'~Spare FB2[273].28'; 8765 '~Spare FB2[273].29'; 8766 '~Spare FB2[273].30'; 8767 '~Spare FB2[273].31'; 8768 '~Spare FB2[274].0'; 8769 '~Spare FB2[274].1'; 8770 '~Spare FB2[274].2'; 8771 '~Spare FB2[274].3'; 8772 '~Spare FB2[274].4'; 8773 '~Spare FB2[274].5'; 8774 '~Spare FB2[274].6'; 8775 '~Spare FB2[274].7'; 8776 '~Spare FB2[274].8'; 8777 '~Spare FB2[274].9'; 8778 '~Spare FB2[274].10'; 8779 '~Spare FB2[274].11'; 8780 '~Spare FB2[274].12'; 8781 '~Spare FB2[274].13'; 8782 '~Spare FB2[274].14'; 8783 '~Spare FB2[274].15'; 8784 '~Spare FB2[274].16'; 8785 '~Spare FB2[274].17'; 8786 '~Spare FB2[274].18'; 8787 '~Spare FB2[274].19'; 8788 '~Spare FB2[274].20'; 8789 '~Spare FB2[274].21'; 8790 '~Spare FB2[274].22'; 8791 '~Spare FB2[274].23'; 8792 '~Spare FB2[274].24'; 8793 '~Spare FB2[274].25'; 8794 '~Spare FB2[274].26'; 8795 '~Spare FB2[274].27'; 8796 '~Spare FB2[274].28'; 8797 '~Spare FB2[274].29'; 8798 '~Spare FB2[274].30'; 8799 '~Spare FB2[274].31'; 8800 '~Spare FB2[275].0'; 8801 '~Spare FB2[275].1'; 8802 '~Spare FB2[275].2'; 8803 '~Spare FB2[275].3'; 8804 '~Spare FB2[275].4'; 8805 '~Spare FB2[275].5'; 8806 '~Spare FB2[275].6'; 8807 '~Spare FB2[275].7'; 8808 '~Spare FB2[275].8'; 8809 '~Spare FB2[275].9'; 8810 '~Spare FB2[275].10'; 8811 '~Spare FB2[275].11'; 8812 '~Spare FB2[275].12'; 8813 '~Spare FB2[275].13'; 8814 '~Spare FB2[275].14'; 8815 '~Spare FB2[275].15'; 8816 '~Spare FB2[275].16'; 8817 '~Spare FB2[275].17'; 8818 '~Spare FB2[275].18'; 8819 '~Spare FB2[275].19'; 8820 '~Spare FB2[275].20'; 8821 '~Spare FB2[275].21'; 8822 '~Spare FB2[275].22'; 8823 '~Spare FB2[275].23'; 8824 '~Spare FB2[275].24'; 8825 '~Spare FB2[275].25'; 8826 '~Spare FB2[275].26'; 8827 '~Spare FB2[275].27'; 8828 '~Spare FB2[275].28'; 8829 '~Spare FB2[275].29'; 8830 '~Spare FB2[275].30'; 8831 '~Spare FB2[275].31'; 8832 '~S001R13CN.I.RbtCtrlFlt - Control Fault FB2[276].0'; 8833 '~S001R13CN.I.CollDetect - Collision Detect FB2[276].1'; 8834 '~S001R13CN.Ix.RbtPromptBox - View Prompt Box at Teach Pendant FB2[276].2'; 8835 '~Spare FB2[276].3'; 8836 '~Spare FB2[276].4'; 8837 '~Spare FB2[276].5'; 8838 '~Spare FB2[276].6'; 8839 '~Spare FB2[276].7'; 8840 '~Spare FB2[276].8'; 8841 '~Spare FB2[276].9'; 8842 '~Spare FB2[276].10'; 8843 '~S001R13CN.I.Wc1WldFlt -Weld Controller 1 Weld Fault FB2[276].11'; 8844 '~S001R13CN.I.Wc1Flt - Weld Timer Flt - Depress Man Weld To Continue FB2[276].12'; 8845 '~S001R13CN.I.Wc1SGunFlt - Weld Controller 1 Servo Gun Fault FB2[276].13'; 8846 '~S001R13CN.I.Wc1SGunMtrTempFlt - Cntrl 1 Servo Gun Motor Over Temp FB2[276].14'; 8847 '~S001R13CN.I.Td1MtrFlt - Tip Dress 1 Motor Fault FB2[276].15'; 8848 '~S001R13CN.I.WC1XfmrTempFlt - Weld Cntrl 1 Transformer Over Temp FB2[276].16'; 8849 '~S001R13CN.I.AutoTipChng1Flt - Auto Tip Changer 1 Fault FB2[276].17'; 8850 '~S001R13CN.I.Slr1NotReady - Seal Controller 1 Not Ready FB2[276].18'; 8851 '~S001R13CN.I.Slr1MajorFlt - Seal Controller 1 Major Fault FB2[276].19'; 8852 '~S001R13CN.I.Slr1VolNotOk - Seal Controller 1 Volume Not Ok Fault FB2[276].20'; 8853 '~S001R13CN.I.Slr1PurgeFlt - Seal Controller 1 Purge Fault FB2[276].21'; 8854 '~S001R13CN.I.Slr1DoserNot Filled - Seal Cntrl 1 Doser Not Filled FB2[276].22'; 8855 '~S001R13CN.I.Slr1No2ClnMxr - Seal Cntrl1 No 2C In Mixer Fault FB2[276].23'; 8856 '~S001R13CN.I.Slr1NzlBroken - Seal Controller 1 Nozzle Broken Fault FB2[276].24'; 8857 '~S001R13CN.I.Slr1NozzleChgReq - Seal Cntrl1 Nozzle Change Reqd FB2[276].25'; 8858 '~S001R13CN.I.Slr1CycleInterrupted - Seal Cntrl1 Cycle Interrupted FB2[276].26'; 8859 '~S001R13CN.I.Stdw1Flt - Stud Weld 1 Weld Fault FB2[276].27'; 8860 '~S001R13CN.I.Stdw1DlyExcdd - Stud Weld 1 Time Delay Exceeded Flt FB2[276].28'; 8861 '~S001R13CN.I.Stdw1Maint Reqd - Stud Weld 1 Maintenance Required FB2[276].29'; 8862 '~S001R13CN.I.Stdw1Reject - Stud Weld 1 art Reject Fault FB2[276].30'; 8863 '~S001R13CN.I.Rvt1Flt - Rivet Controller 1 Fault FB2[276].31'; 8864 '~S001R13CN.I.Rvt1DlyExcdd - Rivet Cntrl 1 Time Delay Exceeded Flt FB2[277].0'; 8865 '~S001R13CN.I.AutoPulledTipByp1 - Auto Pulled Tip Bypass 1 FB2[277].1'; 8866 '~S001R13CN.I.StdWld1EquipmentFlt - Stud Weld 1 Equipment Fault FB2[277].2'; 8867 '~S001R13CN.I.StdWld1BrcktNotPresent - Stud Weld 1 Bracket Not Pres FB2[277].3'; 8868 '~S001R13CN.I.PierceFlt - Pierce Fault FB2[277].4'; 8869 '~S001R13CN.I.NoVisionMeasErr - Vision System Measurement Error FB2[277].5'; 8870 '~S001R13CN.I.VisionSysCalErr - Vision System Calibration Fault FB2[277].6'; 8871 '~S001R13CN.I.VisionSysErr - Vision System Error FB2[277].7'; 8872 '~S001R13CN.I.RackOutOfTolerance - Vision Sys Rack Out Of Tolerance FB2[277].8'; 8873 '~S001R13CN.Ix.TorqFlt - Torque Not Ok FB2[277].9'; 8874 '~S001R13CN.Ix.MwFlt - Mig Weld Controller Fault FB2[277].10'; 8875 '~S001R13CN.Ix.MwWireStuckFlt - Mig Welder Wire Stuck FB2[277].11'; 8876 '~S001R13CN.Ix.MwWldFlt - Mig Welder Bad Bronze Weld Indicator Flt FB2[277].12'; 8877 '~S001R13CN.I.O.TipChngReqd1 - Weld Cntrl 1 Tip Change Required FB2[277].13'; 8878 '~S001R13CN.I.M.NutDetectFlt1 - Nut Welder 1 Nut Detection Fault FB2[277].14'; 8879 '~S001R13CN.I.M.NutProjFlt1 - Nut Welder 1 Weld Not In Tolerance FB2[277].15'; 8880 '~S001R13CN.M.WrongRivetAtNose - Remove Wrong Rivet At Nose FB2[277].16'; 8881 '~S001R13CN.Ix.MwWldLimitErr - Mig Welder CurrentVoltage Out of Tolerance FB2[277].17'; 8882 '~S001R13CN.Ix.MigRdy Mig Welder Not Ready FB2[277].18'; 8883 '~Spare FB2[277].19'; 8884 '~Spare FB2[277].20'; 8885 '~S001R13CN.I.Wc2WldFlt -Weld Controller 2 Weld Fault FB2[277].21'; 8886 '~S001R13CN.I.Wc2Flt - Weld Timer Flt - Depress Man Weld To Continue FB2[277].22'; 8887 '~S001R13CN.I.Wc2SGunFlt - Weld Controller 2 Servo Gun Fault FB2[277].23'; 8888 '~S001R13CN.I.Wc2SGunMtrTempFlt - Cntrl 2 Servo Gun Motor Over Temp FB2[277].24'; 8889 '~S001R13CN.I.Td2MtrFlt - Tip Dress 2 Motor Fault FB2[277].25'; 8890 '~S001R13CN.I.WC2XfmrTempFlt - Weld Cntrl 2 Transformer Over Temp FB2[277].26'; 8891 '~S001R13CN.I.AutoTipChng2Flt - Auto Tip Changer 2 Fault FB2[277].27'; 8892 '~S001R13CN.I.Slr2NotReady - Seal Controller 2 Not Ready FB2[277].28'; 8893 '~S001R13CN.I.Slr2MajorFlt - Seal Controller 2 Major Fault FB2[277].29'; 8894 '~S001R13CN.I.Slr2VolNotOk - Seal Controller 2 Volume Not Ok Fault FB2[277].30'; 8895 '~S001R13CN.I.Slr2PurgeFlt - Seal Controller 2 Purge Fault FB2[277].31'; 8896 '~S001R13CN.I.Slr2DoserNot Filled - Seal Cntrl 2 Doser Not Filled FB2[278].0'; 8897 '~S001R13CN.I.Slr2No2ClnMxr - Seal Cntrl2 No 2C In Mixer Fault FB2[278].1'; 8898 '~S001R13CN.I.Slr2NzlBroken - Seal Controller 2 Nozzle Broken Fault FB2[278].2'; 8899 '~S001R13CN.I.Slr2NozzleChgReq - Seal Cntrl2 Nozzle Change Reqd FB2[278].3'; 8900 '~S001R13CN.I.Slr2CycleInterrupted - Seal Cntrl2 Cycle Interrupted FB2[278].4'; 8901 '~S001R13CN.I.Stdw2Flt - Stud Weld 2 Weld Fault FB2[278].5'; 8902 '~S001R13CN.I.Stdw2DlyExcdd - Stud Weld 2 Time Delay Exceeded Flt FB2[278].6'; 8903 '~S001R13CN.I.Stdw2Maint Reqd - Stud Weld 2 Maintenance Required FB2[278].7'; 8904 '~S001R13CN.I.Stdw2Reject - Stud Weld 2 art Reject Fault FB2[278].8'; 8905 '~S001R13CN.I.Rvt2Flt - Rivet Controller 2 Fault FB2[278].9'; 8906 '~S001R13CN.I.Rvt2DlyExcdd - Rivet Cntrl 2 Time Delay Exceeded Flt FB2[278].10'; 8907 '~S001R13CN.I.AutoPulledTipByp2 - Auto Pulled Tip Bypass 2 FB2[278].11'; 8908 '~S001R13CN.I.StdWld2EquipmentFlt - Stud Weld 2 Equipment Fault FB2[278].12'; 8909 '~S001R13CN.I.StdWld2BrcktNotPresent - Stud Weld 2 Bracket Not Pres FB2[278].13'; 8910 '~S001R13CN.Ix.LsrWldMntrFlt - Seam Geometry/Laser Weld Monitor Flt FB2[278].14'; 8911 '~S001R13CN.Ix.LsrHeadFlt - Laser Head Fault FB2[278].15'; 8912 '~S001R13CN.Ix.LsrGlsFlt - Glass Fault FB2[278].16'; 8913 '~S001R13CN.Ix.LsrWhlFlt - Pressure Wheel Not In Range Fault FB2[278].17'; 8914 '~S001R13CN.Ix.LsrGeoFlt - Seam Geometry/Laser Bad Process Geo Flt FB2[278].18'; 8915 '~S001R13CN.Ix.LsrHdCollFlt - Laser Head Collision Fault FB2[278].19'; 8916 '~S001R13CN.Ix.LsrHdSysFlt - Laser Head System Fault FB2[278].20'; 8917 '~S001R13CN.Ix.LsrHdFar - Laser Head Far Fault FB2[278].21'; 8918 '~S001R13CN.Ix.LsrHdSftCollFlt - Laser Head Software Collision Flt FB2[278].22'; 8919 '~S001R13CN.I.O.TipChngReqd2 - Weld Cntrl 2 Tip Change Required FB2[278].23'; 8920 '~S001R13CN.I.M.NutDetectFlt2 - Nut Welder 2 Nut Detection Fault FB2[278].24'; 8921 '~S001R13CN.I.M.NutProjFlt2 - Nut Welder 2 Weld Not In Tolerance FB2[278].25'; 8922 '~S001R13CN.I.TCWrongToolInStand - Tool Changer Wrong Tool In Stand FB2[278].26'; 8923 '~Spare FB2[278].27'; 8924 '~Spare FB2[278].28'; 8925 '~Spare FB2[278].29'; 8926 '~Spare FB2[278].30'; 8927 '~Spare FB2[278].31'; 8928 '~S001R13CN.I.VisionCommOK - Vision System Comm Fault FB2[279].0'; 8929 '~S001R13CN.I.OutOfTolerance - Vision System Out Of Tolerance FB2[279].1'; 8930 '~S001R13CN.I.MeasureReject - Vision System Measure Reject FB2[279].2'; 8931 '~S001R13CN.I.VisionSysCalibrationFlt - Vision System Calibration Flt FB2[279].3'; 8932 '~S001R13CN.I.VisionSysFlt - Vision System Flt FB2[279].4'; 8933 '~Spare FB2[279].5'; 8934 '~Spare FB2[279].6'; 8935 '~Spare FB2[279].7'; 8936 '~Spare FB2[279].8'; 8937 '~Spare FB2[279].9'; 8938 '~Spare FB2[279].10'; 8939 '~Spare FB2[279].11'; 8940 '~Spare FB2[279].12'; 8941 '~Spare FB2[279].13'; 8942 '~Spare FB2[279].14'; 8943 '~Spare FB2[279].15'; 8944 '~Spare FB2[279].16'; 8945 '~Spare FB2[279].17'; 8946 '~S001R13CN.M.InteruptCyc - Laser Cyc Interupt Cut Wire And Reject Car FB2[279].18'; 8947 '~S001R13CN.M.SuspectPart Inspect Vehicle And Accept Or Reject FB2[279].19'; 8948 '~S001R13 Power Meter High Power Fault Detected FB2[279].20'; 8949 '~S001R13 Power Meter Low Power Fault Detected FB2[279].21'; 8950 '~Spare FB2[279].22'; 8951 '~Spare FB2[279].23'; 8952 '~Spare FB2[279].24'; 8953 '~Spare FB2[279].25'; 8954 '~Spare FB2[279].26'; 8955 '~Spare FB2[279].27'; 8956 '~Spare FB2[279].28'; 8957 '~Spare FB2[279].29'; 8958 '~Spare FB2[279].30'; 8959 '~Spare FB2[279].31'; 8960 '~Spare FB2[280].0'; 8961 '~Spare FB2[280].1'; 8962 '~Spare FB2[280].2'; 8963 '~Spare FB2[280].3'; 8964 '~Spare FB2[280].4'; 8965 '~Spare FB2[280].5'; 8966 '~Spare FB2[280].6'; 8967 '~Spare FB2[280].7'; 8968 '~Spare FB2[280].8'; 8969 '~Spare FB2[280].9'; 8970 '~Spare FB2[280].10'; 8971 '~Spare FB2[280].11'; 8972 '~Spare FB2[280].12'; 8973 '~Spare FB2[280].13'; 8974 '~Spare FB2[280].14'; 8975 '~Spare FB2[280].15'; 8976 '~Spare FB2[280].16'; 8977 '~Spare FB2[280].17'; 8978 '~Spare FB2[280].18'; 8979 '~Spare FB2[280].19'; 8980 '~Spare FB2[280].20'; 8981 '~Spare FB2[280].21'; 8982 '~Spare FB2[280].22'; 8983 '~Spare FB2[280].23'; 8984 '~Spare FB2[280].24'; 8985 '~Spare FB2[280].25'; 8986 '~Spare FB2[280].26'; 8987 '~Spare FB2[280].27'; 8988 '~Spare FB2[280].28'; 8989 '~Spare FB2[280].29'; 8990 '~Spare FB2[280].30'; 8991 '~Spare FB2[280].31'; 8992 '~Spare FB2[281].0'; 8993 '~Spare FB2[281].1'; 8994 '~Spare FB2[281].2'; 8995 '~Spare FB2[281].3'; 8996 '~Spare FB2[281].4'; 8997 '~Spare FB2[281].5'; 8998 '~Spare FB2[281].6'; 8999 '~Spare FB2[281].7'; 9000 '~Spare FB2[281].8'; 9001 '~Spare FB2[281].9'; 9002 '~Spare FB2[281].10'; 9003 '~Spare FB2[281].11'; 9004 '~Spare FB2[281].12'; 9005 '~Spare FB2[281].13'; 9006 '~Spare FB2[281].14'; 9007 '~Spare FB2[281].15'; 9008 '~Spare FB2[281].16'; 9009 '~Spare FB2[281].17'; 9010 '~Spare FB2[281].18'; 9011 '~Spare FB2[281].19'; 9012 '~Spare FB2[281].20'; 9013 '~Spare FB2[281].21'; 9014 '~Spare FB2[281].22'; 9015 '~Spare FB2[281].23'; 9016 '~Spare FB2[281].24'; 9017 '~Spare FB2[281].25'; 9018 '~Spare FB2[281].26'; 9019 '~Spare FB2[281].27'; 9020 '~Spare FB2[281].28'; 9021 '~Spare FB2[281].29'; 9022 '~Spare FB2[281].30'; 9023 '~Spare FB2[281].31'; 9024 '~Spare FB2[282].0'; 9025 '~Spare FB2[282].1'; 9026 '~Spare FB2[282].2'; 9027 '~Spare FB2[282].3'; 9028 '~Spare FB2[282].4'; 9029 '~Spare FB2[282].5'; 9030 '~Spare FB2[282].6'; 9031 '~Spare FB2[282].7'; 9032 '~Spare FB2[282].8'; 9033 '~Spare FB2[282].9'; 9034 '~Spare FB2[282].10'; 9035 '~Spare FB2[282].11'; 9036 '~Spare FB2[282].12'; 9037 '~Spare FB2[282].13'; 9038 '~Spare FB2[282].14'; 9039 '~Spare FB2[282].15'; 9040 '~Spare FB2[282].16'; 9041 '~Spare FB2[282].17'; 9042 '~Spare FB2[282].18'; 9043 '~Spare FB2[282].19'; 9044 '~Spare FB2[282].20'; 9045 '~Spare FB2[282].21'; 9046 '~Spare FB2[282].22'; 9047 '~Spare FB2[282].23'; 9048 '~Spare FB2[282].24'; 9049 '~Spare FB2[282].25'; 9050 '~Spare FB2[282].26'; 9051 '~Spare FB2[282].27'; 9052 '~Spare FB2[282].28'; 9053 '~Spare FB2[282].29'; 9054 '~Spare FB2[282].30'; 9055 '~Spare FB2[282].31'; 9056 '~Spare FB2[283].0'; 9057 '~Spare FB2[283].1'; 9058 '~Spare FB2[283].2'; 9059 '~Spare FB2[283].3'; 9060 '~Spare FB2[283].4'; 9061 '~Spare FB2[283].5'; 9062 '~Spare FB2[283].6'; 9063 '~Spare FB2[283].7'; 9064 '~Spare FB2[283].8'; 9065 '~Spare FB2[283].9'; 9066 '~Spare FB2[283].10'; 9067 '~Spare FB2[283].11'; 9068 '~Spare FB2[283].12'; 9069 '~Spare FB2[283].13'; 9070 '~Spare FB2[283].14'; 9071 '~Spare FB2[283].15'; 9072 '~Spare FB2[283].16'; 9073 '~Spare FB2[283].17'; 9074 '~Spare FB2[283].18'; 9075 '~Spare FB2[283].19'; 9076 '~Spare FB2[283].20'; 9077 '~Spare FB2[283].21'; 9078 '~Spare FB2[283].22'; 9079 '~Spare FB2[283].23'; 9080 '~Spare FB2[283].24'; 9081 '~Spare FB2[283].25'; 9082 '~Spare FB2[283].26'; 9083 '~Spare FB2[283].27'; 9084 '~Spare FB2[283].28'; 9085 '~Spare FB2[283].29'; 9086 '~Spare FB2[283].30'; 9087 '~Spare FB2[283].31'; 9088 '~S001R14CN.I.RbtCtrlFlt - Control Fault FB2[284].0'; 9089 '~S001R14CN.I.CollDetect - Collision Detect FB2[284].1'; 9090 '~S001R14CN.Ix.RbtPromptBox - View Prompt Box at Teach Pendant FB2[284].2'; 9091 '~Spare FB2[284].3'; 9092 '~Spare FB2[284].4'; 9093 '~Spare FB2[284].5'; 9094 '~Spare FB2[284].6'; 9095 '~Spare FB2[284].7'; 9096 '~Spare FB2[284].8'; 9097 '~Spare FB2[284].9'; 9098 '~Spare FB2[284].10'; 9099 '~S001R14CN.I.Wc1WldFlt -Weld Controller 1 Weld Fault FB2[284].11'; 9100 '~S001R14CN.I.Wc1Flt - Weld Timer Flt - Depress Man Weld To Continue FB2[284].12'; 9101 '~S001R14CN.I.Wc1SGunFlt - Weld Controller 1 Servo Gun Fault FB2[284].13'; 9102 '~S001R14CN.I.Wc1SGunMtrTempFlt - Cntrl 1 Servo Gun Motor Over Temp FB2[284].14'; 9103 '~S001R14CN.I.Td1MtrFlt - Tip Dress 1 Motor Fault FB2[284].15'; 9104 '~S001R14CN.I.WC1XfmrTempFlt - Weld Cntrl 1 Transformer Over Temp FB2[284].16'; 9105 '~S001R14CN.I.AutoTipChng1Flt - Auto Tip Changer 1 Fault FB2[284].17'; 9106 '~S001R14CN.I.Slr1NotReady - Seal Controller 1 Not Ready FB2[284].18'; 9107 '~S001R14CN.I.Slr1MajorFlt - Seal Controller 1 Major Fault FB2[284].19'; 9108 '~S001R14CN.I.Slr1VolNotOk - Seal Controller 1 Volume Not Ok Fault FB2[284].20'; 9109 '~S001R14CN.I.Slr1PurgeFlt - Seal Controller 1 Purge Fault FB2[284].21'; 9110 '~S001R14CN.I.Slr1DoserNot Filled - Seal Cntrl 1 Doser Not Filled FB2[284].22'; 9111 '~S001R14CN.I.Slr1No2ClnMxr - Seal Cntrl1 No 2C In Mixer Fault FB2[284].23'; 9112 '~S001R14CN.I.Slr1NzlBroken - Seal Controller 1 Nozzle Broken Fault FB2[284].24'; 9113 '~S001R14CN.I.Slr1NozzleChgReq - Seal Cntrl1 Nozzle Change Reqd FB2[284].25'; 9114 '~S001R14CN.I.Slr1CycleInterrupted - Seal Cntrl1 Cycle Interrupted FB2[284].26'; 9115 '~S001R14CN.I.Stdw1Flt - Stud Weld 1 Weld Fault FB2[284].27'; 9116 '~S001R14CN.I.Stdw1DlyExcdd - Stud Weld 1 Time Delay Exceeded Flt FB2[284].28'; 9117 '~S001R14CN.I.Stdw1Maint Reqd - Stud Weld 1 Maintenance Required FB2[284].29'; 9118 '~S001R14CN.I.Stdw1Reject - Stud Weld 1 art Reject Fault FB2[284].30'; 9119 '~S001R14CN.I.Rvt1Flt - Rivet Controller 1 Fault FB2[284].31'; 9120 '~S001R14CN.I.Rvt1DlyExcdd - Rivet Cntrl 1 Time Delay Exceeded Flt FB2[285].0'; 9121 '~S001R14CN.I.AutoPulledTipByp1 - Auto Pulled Tip Bypass 1 FB2[285].1'; 9122 '~S001R14CN.I.StdWld1EquipmentFlt - Stud Weld 1 Equipment Fault FB2[285].2'; 9123 '~S001R14CN.I.StdWld1BrcktNotPresent - Stud Weld 1 Bracket Not Pres FB2[285].3'; 9124 '~S001R14CN.I.PierceFlt - Pierce Fault FB2[285].4'; 9125 '~S001R14CN.I.NoVisionMeasErr - Vision System Measurement Error FB2[285].5'; 9126 '~S001R14CN.I.VisionSysCalErr - Vision System Calibration Fault FB2[285].6'; 9127 '~S001R14CN.I.VisionSysErr - Vision System Error FB2[285].7'; 9128 '~S001R14CN.I.RackOutOfTolerance - Vision Sys Rack Out Of Tolerance FB2[285].8'; 9129 '~S001R14CN.Ix.TorqFlt - Torque Not Ok FB2[285].9'; 9130 '~S001R14CN.Ix.MwFlt - Mig Weld Controller Fault FB2[285].10'; 9131 '~S001R14CN.Ix.MwWireStuckFlt - Mig Welder Wire Stuck FB2[285].11'; 9132 '~S001R14CN.Ix.MwWldFlt - Mig Welder Bad Bronze Weld Indicator Flt FB2[285].12'; 9133 '~S001R14CN.I.O.TipChngReqd1 - Weld Cntrl 1 Tip Change Required FB2[285].13'; 9134 '~S001R14CN.I.M.NutDetectFlt1 - Nut Welder 1 Nut Detection Fault FB2[285].14'; 9135 '~S001R14CN.I.M.NutProjFlt1 - Nut Welder 1 Weld Not In Tolerance FB2[285].15'; 9136 '~S001R14CN.M.WrongRivetAtNose - Remove Wrong Rivet At Nose FB2[285].16'; 9137 '~S001R14CN.Ix.MwWldLimitErr - Mig Welder CurrentVoltage Out of Tolerance FB2[285].17'; 9138 '~S001R14CN.Ix.MigRdy Mig Welder Not Ready FB2[285].18'; 9139 '~Spare FB2[285].19'; 9140 '~Spare FB2[285].20'; 9141 '~S001R14CN.I.Wc2WldFlt -Weld Controller 2 Weld Fault FB2[285].21'; 9142 '~S001R14CN.I.Wc2Flt - Weld Timer Flt - Depress Man Weld To Continue FB2[285].22'; 9143 '~S001R14CN.I.Wc2SGunFlt - Weld Controller 2 Servo Gun Fault FB2[285].23'; 9144 '~S001R14CN.I.Wc2SGunMtrTempFlt - Cntrl 2 Servo Gun Motor Over Temp FB2[285].24'; 9145 '~S001R14CN.I.Td2MtrFlt - Tip Dress 2 Motor Fault FB2[285].25'; 9146 '~S001R14CN.I.WC2XfmrTempFlt - Weld Cntrl 2 Transformer Over Temp FB2[285].26'; 9147 '~S001R14CN.I.AutoTipChng2Flt - Auto Tip Changer 2 Fault FB2[285].27'; 9148 '~S001R14CN.I.Slr2NotReady - Seal Controller 2 Not Ready FB2[285].28'; 9149 '~S001R14CN.I.Slr2MajorFlt - Seal Controller 2 Major Fault FB2[285].29'; 9150 '~S001R14CN.I.Slr2VolNotOk - Seal Controller 2 Volume Not Ok Fault FB2[285].30'; 9151 '~S001R14CN.I.Slr2PurgeFlt - Seal Controller 2 Purge Fault FB2[285].31'; 9152 '~S001R14CN.I.Slr2DoserNot Filled - Seal Cntrl 2 Doser Not Filled FB2[286].0'; 9153 '~S001R14CN.I.Slr2No2ClnMxr - Seal Cntrl2 No 2C In Mixer Fault FB2[286].1'; 9154 '~S001R14CN.I.Slr2NzlBroken - Seal Controller 2 Nozzle Broken Fault FB2[286].2'; 9155 '~S001R14CN.I.Slr2NozzleChgReq - Seal Cntrl2 Nozzle Change Reqd FB2[286].3'; 9156 '~S001R14CN.I.Slr2CycleInterrupted - Seal Cntrl2 Cycle Interrupted FB2[286].4'; 9157 '~S001R14CN.I.Stdw2Flt - Stud Weld 2 Weld Fault FB2[286].5'; 9158 '~S001R14CN.I.Stdw2DlyExcdd - Stud Weld 2 Time Delay Exceeded Flt FB2[286].6'; 9159 '~S001R14CN.I.Stdw2Maint Reqd - Stud Weld 2 Maintenance Required FB2[286].7'; 9160 '~S001R14CN.I.Stdw2Reject - Stud Weld 2 art Reject Fault FB2[286].8'; 9161 '~S001R14CN.I.Rvt2Flt - Rivet Controller 2 Fault FB2[286].9'; 9162 '~S001R14CN.I.Rvt2DlyExcdd - Rivet Cntrl 2 Time Delay Exceeded Flt FB2[286].10'; 9163 '~S001R14CN.I.AutoPulledTipByp2 - Auto Pulled Tip Bypass 2 FB2[286].11'; 9164 '~S001R14CN.I.StdWld2EquipmentFlt - Stud Weld 2 Equipment Fault FB2[286].12'; 9165 '~S001R14CN.I.StdWld2BrcktNotPresent - Stud Weld 2 Bracket Not Pres FB2[286].13'; 9166 '~S001R14CN.Ix.LsrWldMntrFlt - Seam Geometry/Laser Weld Monitor Flt FB2[286].14'; 9167 '~S001R14CN.Ix.LsrHeadFlt - Laser Head Fault FB2[286].15'; 9168 '~S001R14CN.Ix.LsrGlsFlt - Glass Fault FB2[286].16'; 9169 '~S001R14CN.Ix.LsrWhlFlt - Pressure Wheel Not In Range Fault FB2[286].17'; 9170 '~S001R14CN.Ix.LsrGeoFlt - Seam Geometry/Laser Bad Process Geo Flt FB2[286].18'; 9171 '~S001R14CN.Ix.LsrHdCollFlt - Laser Head Collision Fault FB2[286].19'; 9172 '~S001R14CN.Ix.LsrHdSysFlt - Laser Head System Fault FB2[286].20'; 9173 '~S001R14CN.Ix.LsrHdFar - Laser Head Far Fault FB2[286].21'; 9174 '~S001R14CN.Ix.LsrHdSftCollFlt - Laser Head Software Collision Flt FB2[286].22'; 9175 '~S001R14CN.I.O.TipChngReqd2 - Weld Cntrl 2 Tip Change Required FB2[286].23'; 9176 '~S001R14CN.I.M.NutDetectFlt2 - Nut Welder 2 Nut Detection Fault FB2[286].24'; 9177 '~S001R14CN.I.M.NutProjFlt2 - Nut Welder 2 Weld Not In Tolerance FB2[286].25'; 9178 '~S001R14CN.I.TCWrongToolInStand - Tool Changer Wrong Tool In Stand FB2[286].26'; 9179 '~Spare FB2[286].27'; 9180 '~Spare FB2[286].28'; 9181 '~Spare FB2[286].29'; 9182 '~Spare FB2[286].30'; 9183 '~Spare FB2[286].31'; 9184 '~S001R14CN.I.VisionCommOK - Vision System Comm Fault FB2[287].0'; 9185 '~S001R14CN.I.OutOfTolerance - Vision System Out Of Tolerance FB2[287].1'; 9186 '~S001R14CN.I.MeasureReject - Vision System Measure Reject FB2[287].2'; 9187 '~S001R14CN.I.VisionSysCalibrationFlt - Vision System Calibration Flt FB2[287].3'; 9188 '~S001R14CN.I.VisionSysFlt - Vision System Flt FB2[287].4'; 9189 '~Spare FB2[287].5'; 9190 '~Spare FB2[287].6'; 9191 '~Spare FB2[287].7'; 9192 '~Spare FB2[287].8'; 9193 '~Spare FB2[287].9'; 9194 '~Spare FB2[287].10'; 9195 '~Spare FB2[287].11'; 9196 '~Spare FB2[287].12'; 9197 '~Spare FB2[287].13'; 9198 '~Spare FB2[287].14'; 9199 '~Spare FB2[287].15'; 9200 '~Spare FB2[287].16'; 9201 '~Spare FB2[287].17'; 9202 '~S001R14CN.M.InteruptCyc - Laser Cyc Interupt Cut Wire And Reject Car FB2[287].18'; 9203 '~S001R14CN.M.SuspectPart Inspect Vehicle And Accept Or Reject FB2[287].19'; 9204 '~S001R14 Power Meter High Power Fault Detected FB2[287].20'; 9205 '~S001R14 Power Meter Low Power Fault Detected FB2[287].21'; 9206 '~Spare FB2[287].22'; 9207 '~Spare FB2[287].23'; 9208 '~Spare FB2[287].24'; 9209 '~Spare FB2[287].25'; 9210 '~Spare FB2[287].26'; 9211 '~Spare FB2[287].27'; 9212 '~Spare FB2[287].28'; 9213 '~Spare FB2[287].29'; 9214 '~Spare FB2[287].30'; 9215 '~Spare FB2[287].31'; 9216 '~Spare FB2[288].0'; 9217 '~Spare FB2[288].1'; 9218 '~Spare FB2[288].2'; 9219 '~Spare FB2[288].3'; 9220 '~Spare FB2[288].4'; 9221 '~Spare FB2[288].5'; 9222 '~Spare FB2[288].6'; 9223 '~Spare FB2[288].7'; 9224 '~Spare FB2[288].8'; 9225 '~Spare FB2[288].9'; 9226 '~Spare FB2[288].10'; 9227 '~Spare FB2[288].11'; 9228 '~Spare FB2[288].12'; 9229 '~Spare FB2[288].13'; 9230 '~Spare FB2[288].14'; 9231 '~Spare FB2[288].15'; 9232 '~Spare FB2[288].16'; 9233 '~Spare FB2[288].17'; 9234 '~Spare FB2[288].18'; 9235 '~Spare FB2[288].19'; 9236 '~Spare FB2[288].20'; 9237 '~Spare FB2[288].21'; 9238 '~Spare FB2[288].22'; 9239 '~Spare FB2[288].23'; 9240 '~Spare FB2[288].24'; 9241 '~Spare FB2[288].25'; 9242 '~Spare FB2[288].26'; 9243 '~Spare FB2[288].27'; 9244 '~Spare FB2[288].28'; 9245 '~Spare FB2[288].29'; 9246 '~Spare FB2[288].30'; 9247 '~Spare FB2[288].31'; 9248 '~Spare FB2[289].0'; 9249 '~Spare FB2[289].1'; 9250 '~Spare FB2[289].2'; 9251 '~Spare FB2[289].3'; 9252 '~Spare FB2[289].4'; 9253 '~Spare FB2[289].5'; 9254 '~Spare FB2[289].6'; 9255 '~Spare FB2[289].7'; 9256 '~Spare FB2[289].8'; 9257 '~Spare FB2[289].9'; 9258 '~Spare FB2[289].10'; 9259 '~Spare FB2[289].11'; 9260 '~Spare FB2[289].12'; 9261 '~Spare FB2[289].13'; 9262 '~Spare FB2[289].14'; 9263 '~Spare FB2[289].15'; 9264 '~Spare FB2[289].16'; 9265 '~Spare FB2[289].17'; 9266 '~Spare FB2[289].18'; 9267 '~Spare FB2[289].19'; 9268 '~Spare FB2[289].20'; 9269 '~Spare FB2[289].21'; 9270 '~Spare FB2[289].22'; 9271 '~Spare FB2[289].23'; 9272 '~Spare FB2[289].24'; 9273 '~Spare FB2[289].25'; 9274 '~Spare FB2[289].26'; 9275 '~Spare FB2[289].27'; 9276 '~Spare FB2[289].28'; 9277 '~Spare FB2[289].29'; 9278 '~Spare FB2[289].30'; 9279 '~Spare FB2[289].31'; 9280 '~Spare FB2[290].0'; 9281 '~Spare FB2[290].1'; 9282 '~Spare FB2[290].2'; 9283 '~Spare FB2[290].3'; 9284 '~Spare FB2[290].4'; 9285 '~Spare FB2[290].5'; 9286 '~Spare FB2[290].6'; 9287 '~Spare FB2[290].7'; 9288 '~Spare FB2[290].8'; 9289 '~Spare FB2[290].9'; 9290 '~Spare FB2[290].10'; 9291 '~Spare FB2[290].11'; 9292 '~Spare FB2[290].12'; 9293 '~Spare FB2[290].13'; 9294 '~Spare FB2[290].14'; 9295 '~Spare FB2[290].15'; 9296 '~Spare FB2[290].16'; 9297 '~Spare FB2[290].17'; 9298 '~Spare FB2[290].18'; 9299 '~Spare FB2[290].19'; 9300 '~Spare FB2[290].20'; 9301 '~Spare FB2[290].21'; 9302 '~Spare FB2[290].22'; 9303 '~Spare FB2[290].23'; 9304 '~Spare FB2[290].24'; 9305 '~Spare FB2[290].25'; 9306 '~Spare FB2[290].26'; 9307 '~Spare FB2[290].27'; 9308 '~Spare FB2[290].28'; 9309 '~Spare FB2[290].29'; 9310 '~Spare FB2[290].30'; 9311 '~Spare FB2[290].31'; 9312 '~Spare FB2[291].0'; 9313 '~Spare FB2[291].1'; 9314 '~Spare FB2[291].2'; 9315 '~Spare FB2[291].3'; 9316 '~Spare FB2[291].4'; 9317 '~Spare FB2[291].5'; 9318 '~Spare FB2[291].6'; 9319 '~Spare FB2[291].7'; 9320 '~Spare FB2[291].8'; 9321 '~Spare FB2[291].9'; 9322 '~Spare FB2[291].10'; 9323 '~Spare FB2[291].11'; 9324 '~Spare FB2[291].12'; 9325 '~Spare FB2[291].13'; 9326 '~Spare FB2[291].14'; 9327 '~Spare FB2[291].15'; 9328 '~Spare FB2[291].16'; 9329 '~Spare FB2[291].17'; 9330 '~Spare FB2[291].18'; 9331 '~Spare FB2[291].19'; 9332 '~Spare FB2[291].20'; 9333 '~Spare FB2[291].21'; 9334 '~Spare FB2[291].22'; 9335 '~Spare FB2[291].23'; 9336 '~Spare FB2[291].24'; 9337 '~Spare FB2[291].25'; 9338 '~Spare FB2[291].26'; 9339 '~Spare FB2[291].27'; 9340 '~Spare FB2[291].28'; 9341 '~Spare FB2[291].29'; 9342 '~Spare FB2[291].30'; 9343 '~Spare FB2[291].31'; 9344 '~S001R15CN.I.RbtCtrlFlt - Control Fault FB2[292].0'; 9345 '~S001R15CN.I.CollDetect - Collision Detect FB2[292].1'; 9346 '~S001R15CN.Ix.RbtPromptBox - View Prompt Box at Teach Pendant FB2[292].2'; 9347 '~Spare FB2[292].3'; 9348 '~Spare FB2[292].4'; 9349 '~Spare FB2[292].5'; 9350 '~Spare FB2[292].6'; 9351 '~Spare FB2[292].7'; 9352 '~Spare FB2[292].8'; 9353 '~Spare FB2[292].9'; 9354 '~Spare FB2[292].10'; 9355 '~S001R15CN.I.Wc1WldFlt -Weld Controller 1 Weld Fault FB2[292].11'; 9356 '~S001R15CN.I.Wc1Flt - Weld Timer Flt - Depress Man Weld To Continue FB2[292].12'; 9357 '~S001R15CN.I.Wc1SGunFlt - Weld Controller 1 Servo Gun Fault FB2[292].13'; 9358 '~S001R15CN.I.Wc1SGunMtrTempFlt - Cntrl 1 Servo Gun Motor Over Temp FB2[292].14'; 9359 '~S001R15CN.I.Td1MtrFlt - Tip Dress 1 Motor Fault FB2[292].15'; 9360 '~S001R15CN.I.WC1XfmrTempFlt - Weld Cntrl 1 Transformer Over Temp FB2[292].16'; 9361 '~S001R15CN.I.AutoTipChng1Flt - Auto Tip Changer 1 Fault FB2[292].17'; 9362 '~S001R15CN.I.Slr1NotReady - Seal Controller 1 Not Ready FB2[292].18'; 9363 '~S001R15CN.I.Slr1MajorFlt - Seal Controller 1 Major Fault FB2[292].19'; 9364 '~S001R15CN.I.Slr1VolNotOk - Seal Controller 1 Volume Not Ok Fault FB2[292].20'; 9365 '~S001R15CN.I.Slr1PurgeFlt - Seal Controller 1 Purge Fault FB2[292].21'; 9366 '~S001R15CN.I.Slr1DoserNot Filled - Seal Cntrl 1 Doser Not Filled FB2[292].22'; 9367 '~S001R15CN.I.Slr1No2ClnMxr - Seal Cntrl1 No 2C In Mixer Fault FB2[292].23'; 9368 '~S001R15CN.I.Slr1NzlBroken - Seal Controller 1 Nozzle Broken Fault FB2[292].24'; 9369 '~S001R15CN.I.Slr1NozzleChgReq - Seal Cntrl1 Nozzle Change Reqd FB2[292].25'; 9370 '~S001R15CN.I.Slr1CycleInterrupted - Seal Cntrl1 Cycle Interrupted FB2[292].26'; 9371 '~S001R15CN.I.Stdw1Flt - Stud Weld 1 Weld Fault FB2[292].27'; 9372 '~S001R15CN.I.Stdw1DlyExcdd - Stud Weld 1 Time Delay Exceeded Flt FB2[292].28'; 9373 '~S001R15CN.I.Stdw1Maint Reqd - Stud Weld 1 Maintenance Required FB2[292].29'; 9374 '~S001R15CN.I.Stdw1Reject - Stud Weld 1 art Reject Fault FB2[292].30'; 9375 '~S001R15CN.I.Rvt1Flt - Rivet Controller 1 Fault FB2[292].31'; 9376 '~S001R15CN.I.Rvt1DlyExcdd - Rivet Cntrl 1 Time Delay Exceeded Flt FB2[293].0'; 9377 '~S001R15CN.I.AutoPulledTipByp1 - Auto Pulled Tip Bypass 1 FB2[293].1'; 9378 '~S001R15CN.I.StdWld1EquipmentFlt - Stud Weld 1 Equipment Fault FB2[293].2'; 9379 '~S001R15CN.I.StdWld1BrcktNotPresent - Stud Weld 1 Bracket Not Pres FB2[293].3'; 9380 '~S001R15CN.I.PierceFlt - Pierce Fault FB2[293].4'; 9381 '~S001R15CN.I.NoVisionMeasErr - Vision System Measurement Error FB2[293].5'; 9382 '~S001R15CN.I.VisionSysCalErr - Vision System Calibration Fault FB2[293].6'; 9383 '~S001R15CN.I.VisionSysErr - Vision System Error FB2[293].7'; 9384 '~S001R15CN.I.RackOutOfTolerance - Vision Sys Rack Out Of Tolerance FB2[293].8'; 9385 '~S001R15CN.Ix.TorqFlt - Torque Not Ok FB2[293].9'; 9386 '~S001R15CN.Ix.MwFlt - Mig Weld Controller Fault FB2[293].10'; 9387 '~S001R15CN.Ix.MwWireStuckFlt - Mig Welder Wire Stuck FB2[293].11'; 9388 '~S001R15CN.Ix.MwWldFlt - Mig Welder Bad Bronze Weld Indicator Flt FB2[293].12'; 9389 '~S001R15CN.I.O.TipChngReqd1 - Weld Cntrl 1 Tip Change Required FB2[293].13'; 9390 '~S001R15CN.I.M.NutDetectFlt1 - Nut Welder 1 Nut Detection Fault FB2[293].14'; 9391 '~S001R15CN.I.M.NutProjFlt1 - Nut Welder 1 Weld Not In Tolerance FB2[293].15'; 9392 '~S001R15CN.M.WrongRivetAtNose - Remove Wrong Rivet At Nose FB2[293].16'; 9393 '~S001R15CN.Ix.MwWldLimitErr - Mig Welder CurrentVoltage Out of Tolerance FB2[293].17'; 9394 '~S001R15CN.Ix.MigRdy Mig Welder Not Ready FB2[293].18'; 9395 '~Spare FB2[293].19'; 9396 '~Spare FB2[293].20'; 9397 '~S001R15CN.I.Wc2WldFlt -Weld Controller 2 Weld Fault FB2[293].21'; 9398 '~S001R15CN.I.Wc2Flt - Weld Timer Flt - Depress Man Weld To Continue FB2[293].22'; 9399 '~S001R15CN.I.Wc2SGunFlt - Weld Controller 2 Servo Gun Fault FB2[293].23'; 9400 '~S001R15CN.I.Wc2SGunMtrTempFlt - Cntrl 2 Servo Gun Motor Over Temp FB2[293].24'; 9401 '~S001R15CN.I.Td2MtrFlt - Tip Dress 2 Motor Fault FB2[293].25'; 9402 '~S001R15CN.I.WC2XfmrTempFlt - Weld Cntrl 2 Transformer Over Temp FB2[293].26'; 9403 '~S001R15CN.I.AutoTipChng2Flt - Auto Tip Changer 2 Fault FB2[293].27'; 9404 '~S001R15CN.I.Slr2NotReady - Seal Controller 2 Not Ready FB2[293].28'; 9405 '~S001R15CN.I.Slr2MajorFlt - Seal Controller 2 Major Fault FB2[293].29'; 9406 '~S001R15CN.I.Slr2VolNotOk - Seal Controller 2 Volume Not Ok Fault FB2[293].30'; 9407 '~S001R15CN.I.Slr2PurgeFlt - Seal Controller 2 Purge Fault FB2[293].31'; 9408 '~S001R15CN.I.Slr2DoserNot Filled - Seal Cntrl 2 Doser Not Filled FB2[294].0'; 9409 '~S001R15CN.I.Slr2No2ClnMxr - Seal Cntrl2 No 2C In Mixer Fault FB2[294].1'; 9410 '~S001R15CN.I.Slr2NzlBroken - Seal Controller 2 Nozzle Broken Fault FB2[294].2'; 9411 '~S001R15CN.I.Slr2NozzleChgReq - Seal Cntrl2 Nozzle Change Reqd FB2[294].3'; 9412 '~S001R15CN.I.Slr2CycleInterrupted - Seal Cntrl2 Cycle Interrupted FB2[294].4'; 9413 '~S001R15CN.I.Stdw2Flt - Stud Weld 2 Weld Fault FB2[294].5'; 9414 '~S001R15CN.I.Stdw2DlyExcdd - Stud Weld 2 Time Delay Exceeded Flt FB2[294].6'; 9415 '~S001R15CN.I.Stdw2Maint Reqd - Stud Weld 2 Maintenance Required FB2[294].7'; 9416 '~S001R15CN.I.Stdw2Reject - Stud Weld 2 art Reject Fault FB2[294].8'; 9417 '~S001R15CN.I.Rvt2Flt - Rivet Controller 2 Fault FB2[294].9'; 9418 '~S001R15CN.I.Rvt2DlyExcdd - Rivet Cntrl 2 Time Delay Exceeded Flt FB2[294].10'; 9419 '~S001R15CN.I.AutoPulledTipByp2 - Auto Pulled Tip Bypass 2 FB2[294].11'; 9420 '~S001R15CN.I.StdWld2EquipmentFlt - Stud Weld 2 Equipment Fault FB2[294].12'; 9421 '~S001R15CN.I.StdWld2BrcktNotPresent - Stud Weld 2 Bracket Not Pres FB2[294].13'; 9422 '~S001R15CN.Ix.LsrWldMntrFlt - Seam Geometry/Laser Weld Monitor Flt FB2[294].14'; 9423 '~S001R15CN.Ix.LsrHeadFlt - Laser Head Fault FB2[294].15'; 9424 '~S001R15CN.Ix.LsrGlsFlt - Glass Fault FB2[294].16'; 9425 '~S001R15CN.Ix.LsrWhlFlt - Pressure Wheel Not In Range Fault FB2[294].17'; 9426 '~S001R15CN.Ix.LsrGeoFlt - Seam Geometry/Laser Bad Process Geo Flt FB2[294].18'; 9427 '~S001R15CN.Ix.LsrHdCollFlt - Laser Head Collision Fault FB2[294].19'; 9428 '~S001R15CN.Ix.LsrHdSysFlt - Laser Head System Fault FB2[294].20'; 9429 '~S001R15CN.Ix.LsrHdFar - Laser Head Far Fault FB2[294].21'; 9430 '~S001R15CN.Ix.LsrHdSftCollFlt - Laser Head Software Collision Flt FB2[294].22'; 9431 '~S001R15CN.I.O.TipChngReqd2 - Weld Cntrl 2 Tip Change Required FB2[294].23'; 9432 '~S001R15CN.I.M.NutDetectFlt2 - Nut Welder 2 Nut Detection Fault FB2[294].24'; 9433 '~S001R15CN.I.M.NutProjFlt2 - Nut Welder 2 Weld Not In Tolerance FB2[294].25'; 9434 '~S001R15CN.I.TCWrongToolInStand - Tool Changer Wrong Tool In Stand FB2[294].26'; 9435 '~Spare FB2[294].27'; 9436 '~Spare FB2[294].28'; 9437 '~Spare FB2[294].29'; 9438 '~Spare FB2[294].30'; 9439 '~Spare FB2[294].31'; 9440 '~S001R15CN.I.VisionCommOK - Vision System Comm Fault FB2[295].0'; 9441 '~S001R15CN.I.OutOfTolerance - Vision System Out Of Tolerance FB2[295].1'; 9442 '~S001R15CN.I.MeasureReject - Vision System Measure Reject FB2[295].2'; 9443 '~S001R15CN.I.VisionSysCalibrationFlt - Vision System Calibration Flt FB2[295].3'; 9444 '~S001R15CN.I.VisionSysFlt - Vision System Flt FB2[295].4'; 9445 '~Spare FB2[295].5'; 9446 '~Spare FB2[295].6'; 9447 '~Spare FB2[295].7'; 9448 '~Spare FB2[295].8'; 9449 '~Spare FB2[295].9'; 9450 '~Spare FB2[295].10'; 9451 '~Spare FB2[295].11'; 9452 '~Spare FB2[295].12'; 9453 '~Spare FB2[295].13'; 9454 '~Spare FB2[295].14'; 9455 '~Spare FB2[295].15'; 9456 '~Spare FB2[295].16'; 9457 '~Spare FB2[295].17'; 9458 '~S001R15CN.M.InteruptCyc - Laser Cyc Interupt Cut Wire And Reject Car FB2[295].18'; 9459 '~S001R15CN.M.SuspectPart Inspect Vehicle And Accept Or Reject FB2[295].19'; 9460 '~S001R15 Power Meter High Power Fault Detected FB2[295].20'; 9461 '~S001R15 Power Meter Low Power Fault Detected FB2[295].21'; 9462 '~Spare FB2[295].22'; 9463 '~Spare FB2[295].23'; 9464 '~Spare FB2[295].24'; 9465 '~Spare FB2[295].25'; 9466 '~Spare FB2[295].26'; 9467 '~Spare FB2[295].27'; 9468 '~Spare FB2[295].28'; 9469 '~Spare FB2[295].29'; 9470 '~Spare FB2[295].30'; 9471 '~Spare FB2[295].31'; 9472 '~Spare FB2[296].0'; 9473 '~Spare FB2[296].1'; 9474 '~Spare FB2[296].2'; 9475 '~Spare FB2[296].3'; 9476 '~Spare FB2[296].4'; 9477 '~Spare FB2[296].5'; 9478 '~Spare FB2[296].6'; 9479 '~Spare FB2[296].7'; 9480 '~Spare FB2[296].8'; 9481 '~Spare FB2[296].9'; 9482 '~Spare FB2[296].10'; 9483 '~Spare FB2[296].11'; 9484 '~Spare FB2[296].12'; 9485 '~Spare FB2[296].13'; 9486 '~Spare FB2[296].14'; 9487 '~Spare FB2[296].15'; 9488 '~Spare FB2[296].16'; 9489 '~Spare FB2[296].17'; 9490 '~Spare FB2[296].18'; 9491 '~Spare FB2[296].19'; 9492 '~Spare FB2[296].20'; 9493 '~Spare FB2[296].21'; 9494 '~Spare FB2[296].22'; 9495 '~Spare FB2[296].23'; 9496 '~Spare FB2[296].24'; 9497 '~Spare FB2[296].25'; 9498 '~Spare FB2[296].26'; 9499 '~Spare FB2[296].27'; 9500 '~Spare FB2[296].28'; 9501 '~Spare FB2[296].29'; 9502 '~Spare FB2[296].30'; 9503 '~Spare FB2[296].31'; 9504 '~Spare FB2[297].0'; 9505 '~Spare FB2[297].1'; 9506 '~Spare FB2[297].2'; 9507 '~Spare FB2[297].3'; 9508 '~Spare FB2[297].4'; 9509 '~Spare FB2[297].5'; 9510 '~Spare FB2[297].6'; 9511 '~Spare FB2[297].7'; 9512 '~Spare FB2[297].8'; 9513 '~Spare FB2[297].9'; 9514 '~Spare FB2[297].10'; 9515 '~Spare FB2[297].11'; 9516 '~Spare FB2[297].12'; 9517 '~Spare FB2[297].13'; 9518 '~Spare FB2[297].14'; 9519 '~Spare FB2[297].15'; 9520 '~Spare FB2[297].16'; 9521 '~Spare FB2[297].17'; 9522 '~Spare FB2[297].18'; 9523 '~Spare FB2[297].19'; 9524 '~Spare FB2[297].20'; 9525 '~Spare FB2[297].21'; 9526 '~Spare FB2[297].22'; 9527 '~Spare FB2[297].23'; 9528 '~Spare FB2[297].24'; 9529 '~Spare FB2[297].25'; 9530 '~Spare FB2[297].26'; 9531 '~Spare FB2[297].27'; 9532 '~Spare FB2[297].28'; 9533 '~Spare FB2[297].29'; 9534 '~Spare FB2[297].30'; 9535 '~Spare FB2[297].31'; 9536 '~Spare FB2[298].0'; 9537 '~Spare FB2[298].1'; 9538 '~Spare FB2[298].2'; 9539 '~Spare FB2[298].3'; 9540 '~Spare FB2[298].4'; 9541 '~Spare FB2[298].5'; 9542 '~Spare FB2[298].6'; 9543 '~Spare FB2[298].7'; 9544 '~Spare FB2[298].8'; 9545 '~Spare FB2[298].9'; 9546 '~Spare FB2[298].10'; 9547 '~Spare FB2[298].11'; 9548 '~Spare FB2[298].12'; 9549 '~Spare FB2[298].13'; 9550 '~Spare FB2[298].14'; 9551 '~Spare FB2[298].15'; 9552 '~Spare FB2[298].16'; 9553 '~Spare FB2[298].17'; 9554 '~Spare FB2[298].18'; 9555 '~Spare FB2[298].19'; 9556 '~Spare FB2[298].20'; 9557 '~Spare FB2[298].21'; 9558 '~Spare FB2[298].22'; 9559 '~Spare FB2[298].23'; 9560 '~Spare FB2[298].24'; 9561 '~Spare FB2[298].25'; 9562 '~Spare FB2[298].26'; 9563 '~Spare FB2[298].27'; 9564 '~Spare FB2[298].28'; 9565 '~Spare FB2[298].29'; 9566 '~Spare FB2[298].30'; 9567 '~Spare FB2[298].31'; 9568 '~Spare FB2[299].0'; 9569 '~Spare FB2[299].1'; 9570 '~Spare FB2[299].2'; 9571 '~Spare FB2[299].3'; 9572 '~Spare FB2[299].4'; 9573 '~Spare FB2[299].5'; 9574 '~Spare FB2[299].6'; 9575 '~Spare FB2[299].7'; 9576 '~Spare FB2[299].8'; 9577 '~Spare FB2[299].9'; 9578 '~Spare FB2[299].10'; 9579 '~Spare FB2[299].11'; 9580 '~Spare FB2[299].12'; 9581 '~Spare FB2[299].13'; 9582 '~Spare FB2[299].14'; 9583 '~Spare FB2[299].15'; 9584 '~Spare FB2[299].16'; 9585 '~Spare FB2[299].17'; 9586 '~Spare FB2[299].18'; 9587 '~Spare FB2[299].19'; 9588 '~Spare FB2[299].20'; 9589 '~Spare FB2[299].21'; 9590 '~Spare FB2[299].22'; 9591 '~Spare FB2[299].23'; 9592 '~Spare FB2[299].24'; 9593 '~Spare FB2[299].25'; 9594 '~Spare FB2[299].26'; 9595 '~Spare FB2[299].27'; 9596 '~Spare FB2[299].28'; 9597 '~Spare FB2[299].29'; 9598 '~Spare FB2[299].30'; 9599 '~Spare FB2[299].31'; 9600 '~S001R16CN.I.RbtCtrlFlt - Control Fault FB2[300].0'; 9601 '~S001R16CN.I.CollDetect - Collision Detect FB2[300].1'; 9602 '~S001R16CN.Ix.RbtPromptBox - View Prompt Box at Teach Pendant FB2[300].2'; 9603 '~Spare FB2[300].3'; 9604 '~Spare FB2[300].4'; 9605 '~Spare FB2[300].5'; 9606 '~Spare FB2[300].6'; 9607 '~Spare FB2[300].7'; 9608 '~Spare FB2[300].8'; 9609 '~Spare FB2[300].9'; 9610 '~Spare FB2[300].10'; 9611 '~S001R16CN.I.Wc1WldFlt -Weld Controller 1 Weld Fault FB2[300].11'; 9612 '~S001R16CN.I.Wc1Flt - Weld Timer Flt - Depress Man Weld To Continue FB2[300].12'; 9613 '~S001R16CN.I.Wc1SGunFlt - Weld Controller 1 Servo Gun Fault FB2[300].13'; 9614 '~S001R16CN.I.Wc1SGunMtrTempFlt - Cntrl 1 Servo Gun Motor Over Temp FB2[300].14'; 9615 '~S001R16CN.I.Td1MtrFlt - Tip Dress 1 Motor Fault FB2[300].15'; 9616 '~S001R16CN.I.WC1XfmrTempFlt - Weld Cntrl 1 Transformer Over Temp FB2[300].16'; 9617 '~S001R16CN.I.AutoTipChng1Flt - Auto Tip Changer 1 Fault FB2[300].17'; 9618 '~S001R16CN.I.Slr1NotReady - Seal Controller 1 Not Ready FB2[300].18'; 9619 '~S001R16CN.I.Slr1MajorFlt - Seal Controller 1 Major Fault FB2[300].19'; 9620 '~S001R16CN.I.Slr1VolNotOk - Seal Controller 1 Volume Not Ok Fault FB2[300].20'; 9621 '~S001R16CN.I.Slr1PurgeFlt - Seal Controller 1 Purge Fault FB2[300].21'; 9622 '~S001R16CN.I.Slr1DoserNot Filled - Seal Cntrl 1 Doser Not Filled FB2[300].22'; 9623 '~S001R16CN.I.Slr1No2ClnMxr - Seal Cntrl1 No 2C In Mixer Fault FB2[300].23'; 9624 '~S001R16CN.I.Slr1NzlBroken - Seal Controller 1 Nozzle Broken Fault FB2[300].24'; 9625 '~S001R16CN.I.Slr1NozzleChgReq - Seal Cntrl1 Nozzle Change Reqd FB2[300].25'; 9626 '~S001R16CN.I.Slr1CycleInterrupted - Seal Cntrl1 Cycle Interrupted FB2[300].26'; 9627 '~S001R16CN.I.Stdw1Flt - Stud Weld 1 Weld Fault FB2[300].27'; 9628 '~S001R16CN.I.Stdw1DlyExcdd - Stud Weld 1 Time Delay Exceeded Flt FB2[300].28'; 9629 '~S001R16CN.I.Stdw1Maint Reqd - Stud Weld 1 Maintenance Required FB2[300].29'; 9630 '~S001R16CN.I.Stdw1Reject - Stud Weld 1 art Reject Fault FB2[300].30'; 9631 '~S001R16CN.I.Rvt1Flt - Rivet Controller 1 Fault FB2[300].31'; 9632 '~S001R16CN.I.Rvt1DlyExcdd - Rivet Cntrl 1 Time Delay Exceeded Flt FB2[301].0'; 9633 '~S001R16CN.I.AutoPulledTipByp1 - Auto Pulled Tip Bypass 1 FB2[301].1'; 9634 '~S001R16CN.I.StdWld1EquipmentFlt - Stud Weld 1 Equipment Fault FB2[301].2'; 9635 '~S001R16CN.I.StdWld1BrcktNotPresent - Stud Weld 1 Bracket Not Pres FB2[301].3'; 9636 '~S001R16CN.I.PierceFlt - Pierce Fault FB2[301].4'; 9637 '~S001R16CN.I.NoVisionMeasErr - Vision System Measurement Error FB2[301].5'; 9638 '~S001R16CN.I.VisionSysCalErr - Vision System Calibration Fault FB2[301].6'; 9639 '~S001R16CN.I.VisionSysErr - Vision System Error FB2[301].7'; 9640 '~S001R16CN.I.RackOutOfTolerance - Vision Sys Rack Out Of Tolerance FB2[301].8'; 9641 '~S001R16CN.Ix.TorqFlt - Torque Not Ok FB2[301].9'; 9642 '~S001R16CN.Ix.MwFlt - Mig Weld Controller Fault FB2[301].10'; 9643 '~S001R16CN.Ix.MwWireStuckFlt - Mig Welder Wire Stuck FB2[301].11'; 9644 '~S001R16CN.Ix.MwWldFlt - Mig Welder Bad Bronze Weld Indicator Flt FB2[301].12'; 9645 '~S001R16CN.I.O.TipChngReqd1 - Weld Cntrl 1 Tip Change Required FB2[301].13'; 9646 '~S001R16CN.I.M.NutDetectFlt1 - Nut Welder 1 Nut Detection Fault FB2[301].14'; 9647 '~S001R16CN.I.M.NutProjFlt1 - Nut Welder 1 Weld Not In Tolerance FB2[301].15'; 9648 '~S001R16CN.M.WrongRivetAtNose - Remove Wrong Rivet At Nose FB2[301].16'; 9649 '~S001R16CN.Ix.MwWldLimitErr - Mig Welder CurrentVoltage Out of Tolerance FB2[301].17'; 9650 '~S001R16CN.Ix.MigRdy Mig Welder Not Ready FB2[301].18'; 9651 '~Spare FB2[301].19'; 9652 '~Spare FB2[301].20'; 9653 '~S001R16CN.I.Wc2WldFlt -Weld Controller 2 Weld Fault FB2[301].21'; 9654 '~S001R16CN.I.Wc2Flt - Weld Timer 